                                 END_IF;
                               END_REGION PATH_DYNAMICS

                               REGION CIRCLE_PARAMETERS
                                 IF #statConfigCmdWords[#tempFollowValueCounter].%X4 THEN

                                   // Aux point
                                   FOR #tempCounter := 1 TO 3 DO
                                     IF #statParameterDefinition.followingValues[#tempFollowValueCounter].cmdParameters.circleParameters.auxPoint[#tempCounter] THEN
                                       // Set AuxPoint
                                       #tempParsedValues.cmdParameters.circleParameters.auxPoint[#tempCounter] := #tempParameterValue;
                                       #statParameterValid.cmdParameters.circleParameters.auxPoint[#tempCounter] := TRUE;
                                     END_IF;
                                   END_FOR;

                                   // PathChoice
                                   IF #statParameterDefinition.followingValues[#tempFollowValueCounter].cmdParameters.circleParameters.pathChoice THEN
                                     // Set PathChoice
                                     #tempParsedValues.cmdParameters.circleParameters.pathChoice := LREAL_TO_DINT(#tempParameterValue);
                                     #statParameterValid.cmdParameters.circleParameters.pathChoice := TRUE;
                                   END_IF;


                                   // CircMode
                                   IF #statParameterDefinition.followingValues[#tempFollowValueCounter].cmdParameters.circleParameters.circMode THEN
                                     // Set CircMode
                                     #tempParsedValues.cmdParameters.circleParameters.circMode := LREAL_TO_DINT(#tempParameterValue);
                                     #statParameterValid.cmdParameters.circleParameters.circMode := TRUE;
                                   END_IF;


                                   // CirclePlane
                                   IF #statParameterDefinition.followingValues[#tempFollowValueCounter].cmdParameters.circleParameters.circlePlane THEN
                                     // Set CirclePlane
                                     #tempParsedValues.cmdParameters.circleParameters.circlePlane := LREAL_TO_DINT(#tempParameterValue);
                                     #statParameterValid.cmdParameters.circleParameters.circlePlane := TRUE;
                                   END_IF;


                                   // Arc
                                   IF #statParameterDefinition.followingValues[#tempFollowValueCounter].cmdParameters.circleParameters.arc THEN
                                     // Set Arc
                                     #tempParsedValues.cmdParameters.circleParameters.arc := #tempParameterValue;
                                     #statParameterValid.cmdParameters.circleParameters.arc := TRUE;
                                   END_IF;


                                   // Radius
                                   IF #statParameterDefinition.followingValues[#tempFollowValueCounter].cmdParameters.circleParameters.radius THEN
                                     // Set Radius
                                     #tempParsedValues.cmdParameters.circleParameters.radius := #tempParameterValue;
                                     #statParameterValid.cmdParameters.circleParameters.radius := TRUE;
                                   END_IF;

                                 END_IF;
                               END_REGION CIRCLE_PARAMETERS

                               REGION BOOL_FLAGS
                                 // Always set first index of parsed values here
                                 // ----------------------------------------------------------------------------
                                 // Set Flags
                                 // ----------------------------------------------------------------------------
                                 IF #statParameterDefinition.followingValues[#tempFollowValueCounter].setFlags.flag THEN
                                   // Get parameter value
                                   #tempParsedValues.setFlags[1].flag := LREAL_TO_INT(#tempParameterValue);
                                   #statParameterValid.setFlags[1].flag := TRUE;
                                 END_IF;

                                 // ----------------------------------------------------------------------------
                                 // Flag Mode
                                 // ----------------------------------------------------------------------------
                                 IF #statParameterDefinition.followingValues[#tempFollowValueCounter].setFlags.flagMode THEN
                                   // Get parameter value
                                   #tempParsedValues.setFlags[1].flagMode := LREAL_TO_USINT(#tempParameterValue);
                                   #statParameterValid.setFlags[1].flagMode := TRUE;
                                 END_IF;


                                 // ----------------------------------------------------------------------------
                                 // Remaining Distance
                                 // ----------------------------------------------------------------------------
                                 IF #statParameterDefinition.followingValues[#tempFollowValueCounter].setFlags.remainingDistance THEN
                                   // Get parameter value
                                   #tempParsedValues.setFlags[1].remainingDistance := #tempParameterValue;
                                   #statParameterValid.setFlags[1].remainingDistance := TRUE;
                                 END_IF;

                               END_REGION BOOL_FLAGS

                               REGION LREAL_FLAGS
                                 // Always set first index of parsed values here
                                 // ----------------------------------------------------------------------------
                                 // Set Flags
                                 // ----------------------------------------------------------------------------
                                 IF #statParameterDefinition.followingValues[#tempFollowValueCounter].valueFlags.flag THEN
                                   // Get parameter value
                                   #tempParsedValues.valueFlags[1].flag := LREAL_TO_INT(#tempParameterValue);
                                   #statParameterValid.valueFlags[1].flag := TRUE;
                                 END_IF;

                                 // ----------------------------------------------------------------------------
                                 // Value
                                 // ----------------------------------------------------------------------------
                                 IF #statParameterDefinition.followingValues[#tempFollowValueCounter].valueFlags.value THEN
                                   // Get parameter value
                                   #tempParsedValues.valueFlags[1].value := #tempParameterValue;
                                   #statParameterValid.valueFlags[1].value := TRUE;
                                 END_IF;

                                 // ----------------------------------------------------------------------------
                                 // Flag Mode
                                 // ----------------------------------------------------------------------------
                                 IF #statParameterDefinition.followingValues[#tempFollowValueCounter].valueFlags.flagMode THEN
                                   // Get parameter value
                                   #tempParsedValues.valueFlags[1].flagMode := LREAL_TO_USINT(#tempParameterValue);
                                   #statParameterValid.valueFlags[1].flagMode := TRUE;
                                 END_IF;


                                 // ----------------------------------------------------------------------------
                                 // Remaining Distance
                                 // ----------------------------------------------------------------------------
                                 IF #statParameterDefinition.followingValues[#tempFollowValueCounter].valueFlags.remainingDistance THEN
                                   // Get parameter value
                                   #tempParsedValues.valueFlags[1].remainingDistance := #tempParameterValue;
                                   #statParameterValid.valueFlags[1].remainingDistance := TRUE;
                                 END_IF;

                               END_REGION LREAL_FLAGS

                             END_IF;
                           END_FOR;

                           // Exit loop in case of error
                           IF #statStatus.%X15 THEN
                             EXIT;
                           END_IF;
                         END_REGION GET_FOLLOW_VALUES   
                       END_IF;

                       IF #tempParseCounter = 2 THEN
                         REGION GET_DIRECT_VALUES
                           #tempCmdWord := #statDirectCmdWord;
                           #tempParsedValues := #statParameterDefinition.directValues;
                         END_REGION GET_DIRECT_VALUES
                       END_IF;


                       REGION SET_VALUES_IN_PATH_DATA_ELEMENT

                         IF #tempCmdWord.%X0 THEN

                           REGION CMD_TYPE
                             IF (#statParameterValid.cmdType AND #tempParseCounter = 1)
                               OR (NOT #statParameterValid.cmdType AND #tempParseCounter = 2)
                               AND #statParameterDefinition.priorities.cmdType > "LKINLANG_PRIO_UNRELEVANT"
                             THEN
                               // Get parameter value
                               #tempParameterValue := #tempParsedValues.cmdType;

                               // Set cmdType
                               #statPathDataValue.valueInt := #statActualCommand.pathDataElement.cmdType;
                               #statModalCmdValue.valueInt := #statModalCommand.pathDataElement.cmdType;
                               #statModalPrgValue.valueInt := #statModalProgram.pathDataElement.cmdType;

                               // Set value with follow val from above 
                               #tempReturnVal := "LKinLang_SetValue"(parameterValue := #tempParameterValue,
                                                                     parameterPriority := #statParameterDefinition.priorities.cmdType,
                                                                     validCountOfParameter := #statValidCounts.cmdType,
                                                                     parameterValueMin := -1,
                                                                     parameterValueMax := 100,
                                                                     properties := #statParameterDefinition.properties,
                                                                     errorString => #statErrorString,
                                                                     parameterCounter := #statElementCounter.cmdType,
                                                                     priorityCounter := #statActualCommand.priority.cmdType,
                                                                     modalCMDPrio := #statModalCommand.priority.cmdType,
                                                                     modalPRGPrio := #statModalProgram.priority.cmdType,
                                                                     parameterCounterInLine := #statElementCounterInLine.cmdType,
                                                                     pathDataValue := #statPathDataValue,
                                                                     modalCMDPathDataValue := #statModalCmdValue,
                                                                     modalPRGPathDataValue := #statModalPrgValue);

                               IF #tempReturnVal = 0 THEN
                                 #statActualCommand.pathDataElement.cmdType := #statPathDataValue.valueInt;
                                 #statModalCommand.pathDataElement.cmdType := #statModalCmdValue.valueInt;
                                 #statModalProgram.pathDataElement.cmdType := #statModalPrgValue.valueInt;
                               ELSE
                                 // Error
                                 #statStatus := #ERR_PARSING;
                                 #statErrorString := CONCAT(IN1 := #statErrorString, IN2 := '; Line: ');
                                 #statErrorString := CONCAT(IN1 := #statErrorString, IN2 := UDINT_TO_STRING(#statTokenizedLine.lineNo));
                                 EXIT;
                               END_IF;
                             END_IF;
                           END_REGION CMD_TYPE

                           REGION CMD_NAME
                             IF ((#statParameterValid.cmdName AND #tempParseCounter = 1)
                               OR (NOT #statParameterValid.cmdName AND #tempParseCounter = 2))
                               AND #tempParsedValues.cmdName <> ''
                               AND #statParameterDefinition.priorities.cmdName > "LKINLANG_PRIO_UNRELEVANT"
                             THEN

                               // Get parameter value
                               #tempParameterValue := STRING_TO_INT(#tempParsedValues.cmdName);

                               // Set cmdName
                               #statPathDataValue.valueInt := STRING_TO_INT(#statActualCommand.pathDataElement.cmdName);
                               #statModalCmdValue.valueInt := STRING_TO_INT(#statModalCommand.pathDataElement.cmdName);
                               #statModalPrgValue.valueInt := STRING_TO_INT(#statModalProgram.pathDataElement.cmdName);

                               // Set value with follow val from above 
                               #tempReturnVal := "LKinLang_SetValue"(parameterValue := #tempParameterValue,
                                                                     parameterPriority := #statParameterDefinition.priorities.cmdName,
                                                                     validCountOfParameter := #statValidCounts.cmdName,
                                                                     parameterValueMin := #MINVAL_INT,
                                                                     parameterValueMax := #MAXVAL_INT,
                                                                     properties := #statParameterDefinition.properties,
                                                                     errorString => #statErrorString,
                                                                     parameterCounter := #statElementCounter.cmdName,
                                                                     priorityCounter := #statActualCommand.priority.cmdName,
                                                                     modalCMDPrio := #statModalCommand.priority.cmdName,
                                                                     modalPRGPrio := #statModalProgram.priority.cmdName,
                                                                     parameterCounterInLine := #statElementCounterInLine.cmdName,
                                                                     pathDataValue := #statPathDataValue,
                                                                     modalCMDPathDataValue := #statModalCmdValue,
                                                                     modalPRGPathDataValue := #statModalPrgValue);

                               IF #tempReturnVal = 0 THEN
                                 #statActualCommand.pathDataElement.cmdName := INT_TO_STRING(#statPathDataValue.valueInt);

                                 // 16.07.2019 FR: Delete "+" sign from string
                                 IF #statPathDataValue.valueInt >= 0.0 THEN
                                   #statActualCommand.pathDataElement.cmdName := DELETE(IN := #statActualCommand.pathDataElement.cmdName, L := 1, P := 1);
                                 ELSE
                                   ; // Keep "-" sign
                                 END_IF;

                                 #statModalCommand.pathDataElement.cmdName := INT_TO_STRING(#statModalCmdValue.valueInt);
                                 #statModalProgram.pathDataElement.cmdName := INT_TO_STRING(#statModalPrgValue.valueInt);
                               ELSE
                                 // Error
                                 #statStatus := #ERR_PARSING;
                                 #statErrorString := CONCAT(IN1 := #statErrorString, IN2 := '; Line: ');
                                 #statErrorString := CONCAT(IN1 := #statErrorString, IN2 := UDINT_TO_STRING(#statTokenizedLine.lineNo));
                                 EXIT;
                               END_IF;
                             END_IF;
                           END_REGION CMD_NAME

                           REGION COORDINATES
                             IF #tempCmdWord.%X1 THEN // Coordinates are set

                               // X coordinate
                               IF (#statParameterValid.cmdCoordinates.cartesianPosition.x AND #tempParseCounter = 1)
                                 OR (NOT #statParameterValid.cmdCoordinates.cartesianPosition.x AND #tempParseCounter = 2)
                                 AND #statParameterDefinition.priorities.cmdCoordinates.cartesianPosition.x > "LKINLANG_PRIO_UNRELEVANT"
                               THEN

                                 // Get parameter value
                                 #tempParameterValue := #tempParsedValues.cmdCoordinates.cartesianPosition.x;

                                 // Set X
                                 #statPathDataValue.valueLReal := #statActualCommand.pathDataElement.cmdCoordinates.cartesianPosition.x;
                                 #statModalCmdValue.valueLReal := #statModalCommand.pathDataElement.cmdCoordinates.cartesianPosition.x;
                                 #statModalPrgValue.valueLReal := #statModalProgram.pathDataElement.cmdCoordinates.cartesianPosition.x;

                                 // Set value with follow val from above 
                                 #tempReturnVal := "LKinLang_SetValue"(parameterValue := #tempParameterValue,
                                                                       parameterPriority := #statParameterDefinition.priorities.cmdCoordinates.cartesianPosition.x,
                                                                       validCountOfParameter := #statValidCounts.cmdCoordinates.cartesianPosition.x,
                                                                       parameterValueMin := #MINVAL_LREAL,
                                                                       parameterValueMax := #MAXVAL_LREAL,
                                                                       properties := #statParameterDefinition.properties,
                                                                       errorString => #statErrorString,
                                                                       parameterCounter := #statElementCounter.cmdCoordinates.cartesianPosition.x,
                                                                       priorityCounter := #statActualCommand.priority.cmdCoordinates.cartesianPosition.x,
                                                                       modalCMDPrio := #statModalCommand.priority.cmdCoordinates.cartesianPosition.x,
                                                                       modalPRGPrio := #statModalProgram.priority.cmdCoordinates.cartesianPosition.x,
                                                                       parameterCounterInLine := #statElementCounterInLine.cmdCoordinates.cartesianPosition.x,
                                                                       pathDataValue := #statPathDataValue,
                                                                       modalCMDPathDataValue := #statModalCmdValue,
                                                                       modalPRGPathDataValue := #statModalPrgValue);

                                 IF #tempReturnVal = 0 THEN
                                   #statActualCommand.pathDataElement.cmdCoordinates.cartesianPosition.x := #statPathDataValue.valueLReal;
                                   #statModalCommand.pathDataElement.cmdCoordinates.cartesianPosition.x := #statModalCmdValue.valueLReal;
                                   #statModalProgram.pathDataElement.cmdCoordinates.cartesianPosition.x := #statModalPrgValue.valueLReal;

                                   // Set parameter valid bit for MovePath 
                                   #statActualCommand.pathDataElement.parameterValid[1] := TRUE;
                                 ELSE
                                   // Error
                                   #statStatus := #ERR_PARSING;
                                   #statErrorString := CONCAT(IN1 := #statErrorString, IN2 := '; Line: ');
                                   #statErrorString := CONCAT(IN1 := #statErrorString, IN2 := UDINT_TO_STRING(#statTokenizedLine.lineNo));
                                   EXIT;
                                 END_IF;
                               END_IF;


                               // Y coordinate
                               IF (#statParameterValid.cmdCoordinates.cartesianPosition.y AND #tempParseCounter = 1)
                                 OR (NOT #statParameterValid.cmdCoordinates.cartesianPosition.y AND #tempParseCounter = 2)
                                 AND #statParameterDefinition.priorities.cmdCoordinates.cartesianPosition.y > "LKINLANG_PRIO_UNRELEVANT"
                               THEN

                                 // Get parameter value
                                 #tempParameterValue := #tempParsedValues.cmdCoordinates.cartesianPosition.y;

                                 // Set Y
                                 #statPathDataValue.valueLReal := #statActualCommand.pathDataElement.cmdCoordinates.cartesianPosition.y;
                                 #statModalCmdValue.valueLReal := #statModalCommand.pathDataElement.cmdCoordinates.cartesianPosition.y;
                                 #statModalPrgValue.valueLReal := #statModalProgram.pathDataElement.cmdCoordinates.cartesianPosition.y;

                                 // Set value with follow val from above 
                                 #tempReturnVal := "LKinLang_SetValue"(parameterValue := #tempParameterValue,
                                                                       parameterPriority := #statParameterDefinition.priorities.cmdCoordinates.cartesianPosition.y,
                                                                       validCountOfParameter := #statValidCounts.cmdCoordinates.cartesianPosition.y,
                                                                       parameterValueMin := #MINVAL_LREAL,
                                                                       parameterValueMax := #MAXVAL_LREAL,
                                                                       properties := #statParameterDefinition.properties,
                                                                       errorString => #statErrorString,
                                                                       parameterCounter := #statElementCounter.cmdCoordinates.cartesianPosition.y,
                                                                       priorityCounter := #statActualCommand.priority.cmdCoordinates.cartesianPosition.y,
                                                                       modalCMDPrio := #statModalCommand.priority.cmdCoordinates.cartesianPosition.y,
                                                                       modalPRGPrio := #statModalProgram.priority.cmdCoordinates.cartesianPosition.y,
                                                                       parameterCounterInLine := #statElementCounterInLine.cmdCoordinates.cartesianPosition.y,
                                                                       pathDataValue := #statPathDataValue,
                                                                       modalCMDPathDataValue := #statModalCmdValue,
                                                                       modalPRGPathDataValue := #statModalPrgValue);

                                 IF #tempReturnVal = 0 THEN
                                   #statActualCommand.pathDataElement.cmdCoordinates.cartesianPosition.y := #statPathDataValue.valueLReal;
                                   #statModalCommand.pathDataElement.cmdCoordinates.cartesianPosition.y := #statModalCmdValue.valueLReal;
                                   #statModalProgram.pathDataElement.cmdCoordinates.cartesianPosition.y := #statModalPrgValue.valueLReal;

                                   // Set parameter valid bit for MovePath 
                                   #statActualCommand.pathDataElement.parameterValid[2] := TRUE;
                                 ELSE
                                   // Error
                                   #statStatus := #ERR_PARSING;
                                   #statErrorString := CONCAT(IN1 := #statErrorString, IN2 := '; Line: ');
                                   #statErrorString := CONCAT(IN1 := #statErrorString, IN2 := UDINT_TO_STRING(#statTokenizedLine.lineNo));
                                   EXIT;
                                 END_IF;
                               END_IF;



                               // Z coordinate
                               IF (#statParameterValid.cmdCoordinates.cartesianPosition.z AND #tempParseCounter = 1)
                                 OR (NOT #statParameterValid.cmdCoordinates.cartesianPosition.z AND #tempParseCounter = 2)
                                 AND #statParameterDefinition.priorities.cmdCoordinates.cartesianPosition.z > "LKINLANG_PRIO_UNRELEVANT"
                               THEN

                                 // Get parameter value
                                 #tempParameterValue := #tempParsedValues.cmdCoordinates.cartesianPosition.z;

                                 // Set Z
                                 #statPathDataValue.valueLReal := #statActualCommand.pathDataElement.cmdCoordinates.cartesianPosition.z;
                                 #statModalCmdValue.valueLReal := #statModalCommand.pathDataElement.cmdCoordinates.cartesianPosition.z;
                                 #statModalPrgValue.valueLReal := #statModalProgram.pathDataElement.cmdCoordinates.cartesianPosition.z;

                                 // Set value with follow val from above 
                                 #tempReturnVal := "LKinLang_SetValue"(parameterValue := #tempParameterValue,
                                                                       parameterPriority := #statParameterDefinition.priorities.cmdCoordinates.cartesianPosition.z,
                                                                       validCountOfParameter := #statValidCounts.cmdCoordinates.cartesianPosition.z,
                                                                       parameterValueMin := #MINVAL_LREAL,
                                                                       parameterValueMax := #MAXVAL_LREAL,
                                                                       properties := #statParameterDefinition.properties,
                                                                       errorString => #statErrorString,
                                                                       parameterCounter := #statElementCounter.cmdCoordinates.cartesianPosition.z,
                                                                       priorityCounter := #statActualCommand.priority.cmdCoordinates.cartesianPosition.z,
                                                                       modalCMDPrio := #statModalCommand.priority.cmdCoordinates.cartesianPosition.z,
                                                                       modalPRGPrio := #statModalProgram.priority.cmdCoordinates.cartesianPosition.z,
                                                                       parameterCounterInLine := #statElementCounterInLine.cmdCoordinates.cartesianPosition.z,
                                                                       pathDataValue := #statPathDataValue,
                                                                       modalCMDPathDataValue := #statModalCmdValue,
                                                                       modalPRGPathDataValue := #statModalPrgValue);

                                 IF #tempReturnVal = 0 THEN
                                   #statActualCommand.pathDataElement.cmdCoordinates.cartesianPosition.z := #statPathDataValue.valueLReal;
                                   #statModalCommand.pathDataElement.cmdCoordinates.cartesianPosition.z := #statModalCmdValue.valueLReal;
                                   #statModalProgram.pathDataElement.cmdCoordinates.cartesianPosition.z := #statModalPrgValue.valueLReal;

                                   // Set parameter valid bit for MovePath 
                                   #statActualCommand.pathDataElement.parameterValid[3] := TRUE;
                                 ELSE
                                   // Error
                                   #statStatus := #ERR_PARSING;
                                   #statErrorString := CONCAT(IN1 := #statErrorString, IN2 := '; Line: ');
                                   #statErrorString := CONCAT(IN1 := #statErrorString, IN2 := UDINT_TO_STRING(#statTokenizedLine.lineNo));
                                   EXIT;
                                 END_IF;
                               END_IF;


                               // A coordinate
                               IF (#statParameterValid.cmdCoordinates.cartesianPosition.a AND #tempParseCounter = 1)
                                 OR (NOT #statParameterValid.cmdCoordinates.cartesianPosition.a AND #tempParseCounter = 2)
                                 AND #statParameterDefinition.priorities.cmdCoordinates.cartesianPosition.a > "LKINLANG_PRIO_UNRELEVANT"
                               THEN

                                 // Get parameter value
                                 #tempParameterValue := #tempParsedValues.cmdCoordinates.cartesianPosition.a;

                                 // Set A
                                 #statPathDataValue.valueLReal := #statActualCommand.pathDataElement.cmdCoordinates.cartesianPosition.a;
                                 #statModalCmdValue.valueLReal := #statModalCommand.pathDataElement.cmdCoordinates.cartesianPosition.a;
                                 #statModalPrgValue.valueLReal := #statModalProgram.pathDataElement.cmdCoordinates.cartesianPosition.a;

                                 // Set value with follow val from above 
                                 #tempReturnVal := "LKinLang_SetValue"(parameterValue := #tempParameterValue,
                                                                       parameterPriority := #statParameterDefinition.priorities.cmdCoordinates.cartesianPosition.a,
                                                                       validCountOfParameter := #statValidCounts.cmdCoordinates.cartesianPosition.a,
                                                                       parameterValueMin := #MINVAL_LREAL,
                                                                       parameterValueMax := #MAXVAL_LREAL,
                                                                       properties := #statParameterDefinition.properties,
                                                                       errorString => #statErrorString,
                                                                       parameterCounter := #statElementCounter.cmdCoordinates.cartesianPosition.a,
                                                                       priorityCounter := #statActualCommand.priority.cmdCoordinates.cartesianPosition.a,
                                                                       modalCMDPrio := #statModalCommand.priority.cmdCoordinates.cartesianPosition.a,
                                                                       modalPRGPrio := #statModalProgram.priority.cmdCoordinates.cartesianPosition.a,
                                                                       parameterCounterInLine := #statElementCounterInLine.cmdCoordinates.cartesianPosition.a,
                                                                       pathDataValue := #statPathDataValue,
                                                                       modalCMDPathDataValue := #statModalCmdValue,
                                                                       modalPRGPathDataValue := #statModalPrgValue);

                                 IF #tempReturnVal = 0 THEN
                                   #statActualCommand.pathDataElement.cmdCoordinates.cartesianPosition.a := #statPathDataValue.valueLReal;
                                   #statModalCommand.pathDataElement.cmdCoordinates.cartesianPosition.a := #statModalCmdValue.valueLReal;
                                   #statModalProgram.pathDataElement.cmdCoordinates.cartesianPosition.a := #statModalPrgValue.valueLReal;

                                   // Set parameter valid bit for MovePath 
                                   #statActualCommand.pathDataElement.parameterValid[4] := TRUE;
                                 ELSE
                                   // Error
                                   #statStatus := #ERR_PARSING;
                                   #statErrorString := CONCAT(IN1 := #statErrorString, IN2 := '; Line: ');
                                   #statErrorString := CONCAT(IN1 := #statErrorString, IN2 := UDINT_TO_STRING(#statTokenizedLine.lineNo));
                                   EXIT;
                                 END_IF;
                               END_IF;


                               // CoordSystem coordinate
                               IF (#statParameterValid.cmdCoordinates.coordSystem AND #tempParseCounter = 1)
                                 OR (NOT #statParameterValid.cmdCoordinates.coordSystem AND #tempParseCounter = 2)
                                 AND #statParameterDefinition.priorities.cmdCoordinates.coordSystem > "LKINLANG_PRIO_UNRELEVANT"
                               THEN

                                 // Get parameter value
                                 #tempParameterValue := #tempParsedValues.cmdCoordinates.coordSystem;

                                 // Set CS
                                 #statPathDataValue.valueDint := #statActualCommand.pathDataElement.cmdCoordinates.coordSystem;
                                 #statModalCmdValue.valueDint := #statModalCommand.pathDataElement.cmdCoordinates.coordSystem;
                                 #statModalPrgValue.valueDint := #statModalProgram.pathDataElement.cmdCoordinates.coordSystem;

                                 // Set value with follow val from above 
                                 #tempReturnVal := "LKinLang_SetValue"(parameterValue := #tempParameterValue,
                                                                       parameterPriority := #statParameterDefinition.priorities.cmdCoordinates.coordSystem,
                                                                       validCountOfParameter := #statValidCounts.cmdCoordinates.coordSystem,
                                                                       parameterValueMin := 0,
                                                                       parameterValueMax := 3,
                                                                       properties := #statParameterDefinition.properties,
                                                                       errorString => #statErrorString,
                                                                       parameterCounter := #statElementCounter.cmdCoordinates.coordSystem,
                                                                       priorityCounter := #statActualCommand.priority.cmdCoordinates.coordSystem,
                                                                       modalCMDPrio := #statModalCommand.priority.cmdCoordinates.coordSystem,
                                                                       modalPRGPrio := #statModalProgram.priority.cmdCoordinates.coordSystem,
                                                                       parameterCounterInLine := #statElementCounterInLine.cmdCoordinates.coordSystem,
                                                                       pathDataValue := #statPathDataValue,
                                                                       modalCMDPathDataValue := #statModalCmdValue,
                                                                       modalPRGPathDataValue := #statModalPrgValue);

                                 IF #tempReturnVal = 0 THEN
                                   #statActualCommand.pathDataElement.cmdCoordinates.coordSystem := #statPathDataValue.valueDint;
                                   #statModalCommand.pathDataElement.cmdCoordinates.coordSystem := #statModalCmdValue.valueDint;
                                   #statModalProgram.pathDataElement.cmdCoordinates.coordSystem := #statModalPrgValue.valueDint;
                                 ELSE
                                   // Error
                                   #statStatus := #ERR_PARSING;
                                   #statErrorString := CONCAT(IN1 := #statErrorString, IN2 := '; Line: ');
                                   #statErrorString := CONCAT(IN1 := #statErrorString, IN2 := UDINT_TO_STRING(#statTokenizedLine.lineNo));
                                   EXIT;
                                 END_IF;
                               END_IF;

                             END_IF;
                           END_REGION COORDINATES

                           REGION CMD_PARAMETERS

                             IF #tempCmdWord.%X2 THEN // Parameter are to be set

                               REGION GENERAL_PARAMETERS

                                 // Buffer mode
                                 IF (#statParameterValid.cmdParameters.bufferMode AND #tempParseCounter = 1)
                                   OR (NOT #statParameterValid.cmdParameters.bufferMode AND #tempParseCounter = 2)
                                   AND #statParameterDefinition.priorities.cmdParameters.bufferMode > "LKINLANG_PRIO_UNRELEVANT"
                                 THEN

                                   // Get parameter value
                                   #tempParameterValue := #tempParsedValues.cmdParameters.bufferMode;

                                   // Set Velocity
                                   #statPathDataValue.valueDint := #statActualCommand.pathDataElement.cmdParameters.bufferMode;
                                   #statModalCmdValue.valueDint := #statModalCommand.pathDataElement.cmdParameters.bufferMode;
                                   #statModalPrgValue.valueDint := #statModalProgram.pathDataElement.cmdParameters.bufferMode;

                                   // Set value with follow val from above 
                                   #tempReturnVal := "LKinLang_SetValue"(parameterValue := #tempParameterValue,
                                                                         parameterPriority := #statParameterDefinition.priorities.cmdParameters.bufferMode,
                                                                         validCountOfParameter := #statValidCounts.cmdParameters.bufferMode,
                                                                         parameterValueMin := 1,
                                                                         parameterValueMax := 5,
                                                                         properties := #statParameterDefinition.properties,
                                                                         errorString => #statErrorString,
                                                                         parameterCounter := #statElementCounter.cmdParameters.bufferMode,
                                                                         priorityCounter := #statActualCommand.priority.cmdParameters.bufferMode,
                                                                         modalCMDPrio := #statModalCommand.priority.cmdParameters.bufferMode,
                                                                         modalPRGPrio := #statModalProgram.priority.cmdParameters.bufferMode,
                                                                         parameterCounterInLine := #statElementCounterInLine.cmdParameters.bufferMode,
                                                                         pathDataValue := #statPathDataValue,
                                                                         modalCMDPathDataValue := #statModalCmdValue,
                                                                         modalPRGPathDataValue := #statModalPrgValue);

                                   IF #tempReturnVal = 0 THEN
                                     #statActualCommand.pathDataElement.cmdParameters.bufferMode := #statPathDataValue.valueDint;
                                     #statModalCommand.pathDataElement.cmdParameters.bufferMode := #statModalCmdValue.valueDint;
                                     #statModalProgram.pathDataElement.cmdParameters.bufferMode := #statModalPrgValue.valueDint;
                                   ELSE
                                     // Error
                                     #statStatus := #ERR_PARSING;
                                     #statErrorString := CONCAT(IN1 := #statErrorString, IN2 := '; Line: ');
                                     #statErrorString := CONCAT(IN1 := #statErrorString, IN2 := UDINT_TO_STRING(#statTokenizedLine.lineNo));
                                     EXIT;
                                   END_IF;
                                 END_IF;

                                 // Dynamic adaption
                                 IF (#statParameterValid.cmdParameters.dynamicAdaption AND #tempParseCounter = 1)
                                   OR (NOT #statParameterValid.cmdParameters.dynamicAdaption AND #tempParseCounter = 2)
                                   AND #statParameterDefinition.priorities.cmdParameters.dynamicAdaption > "LKINLANG_PRIO_UNRELEVANT"
                                 THEN

                                   // Get parameter value
                                   #tempParameterValue := #tempParsedValues.cmdParameters.dynamicAdaption;

                                   // Set Velocity
                                   #statPathDataValue.valueDint := #statActualCommand.pathDataElement.cmdParameters.dynamicAdaption;
                                   #statModalCmdValue.valueDint := #statModalCommand.pathDataElement.cmdParameters.dynamicAdaption;
                                   #statModalPrgValue.valueDint := #statModalProgram.pathDataElement.cmdParameters.dynamicAdaption;

                                   // Set value with follow val from above 
                                   #tempReturnVal := "LKinLang_SetValue"(parameterValue := #tempParameterValue,
                                                                         parameterPriority := #statParameterDefinition.priorities.cmdParameters.dynamicAdaption,
                                                                         validCountOfParameter := #statValidCounts.cmdParameters.dynamicAdaption,
                                                                         parameterValueMin := -1,
                                                                         parameterValueMax := 2,
                                                                         properties := #statParameterDefinition.properties,
                                                                         errorString => #statErrorString,
                                                                         parameterCounter := #statElementCounter.cmdParameters.dynamicAdaption,
                                                                         priorityCounter := #statActualCommand.priority.cmdParameters.dynamicAdaption,
                                                                         modalCMDPrio := #statModalCommand.priority.cmdParameters.dynamicAdaption,
                                                                         modalPRGPrio := #statModalProgram.priority.cmdParameters.dynamicAdaption,
                                                                         parameterCounterInLine := #statElementCounterInLine.cmdParameters.dynamicAdaption,
                                                                         pathDataValue := #statPathDataValue,
                                                                         modalCMDPathDataValue := #statModalCmdValue,
                                                                         modalPRGPathDataValue := #statModalPrgValue);

                                   IF #tempReturnVal = 0 THEN
                                     #statActualCommand.pathDataElement.cmdParameters.dynamicAdaption := #statPathDataValue.valueDint;
                                     #statModalCommand.pathDataElement.cmdParameters.dynamicAdaption := #statModalCmdValue.valueDint;
                                     #statModalProgram.pathDataElement.cmdParameters.dynamicAdaption := #statModalPrgValue.valueDint;
                                   ELSE
                                     // Error
                                     #statStatus := #ERR_PARSING;
                                     #statErrorString := CONCAT(IN1 := #statErrorString, IN2 := '; Line: ');
                                     #statErrorString := CONCAT(IN1 := #statErrorString, IN2 := UDINT_TO_STRING(#statTokenizedLine.lineNo));
                                     EXIT;
                                   END_IF;
                                 END_IF;

                                 // Offset Parameter
                                 // Offset Parameter number
                                 IF (#statParameterValid.cmdParameters.offsetParameters.offsetParaNo AND #tempParseCounter = 1)
                                   OR (NOT #statParameterValid.cmdParameters.offsetParameters.offsetParaNo AND #tempParseCounter = 2)
                                   AND #statParameterDefinition.priorities.cmdParameters.offsetParameters.offsetParaNo > "LKINLANG_PRIO_UNRELEVANT"
                                 THEN

                                   // Get parameter value
                                   #tempParameterValue := #tempParsedValues.cmdParameters.offsetParameters.offsetParaNo;

                                   // Set Velocity
                                   #statPathDataValue.valueDint := #statActualCommand.pathDataElement.cmdParameters.offsetParameters.offsetParaNo;
                                   #statModalCmdValue.valueDint := #statModalCommand.pathDataElement.cmdParameters.offsetParameters.offsetParaNo;
                                   #statModalPrgValue.valueDint := #statModalProgram.pathDataElement.cmdParameters.offsetParameters.offsetParaNo;

                                   // Set value with follow val from above 
                                   #tempReturnVal := "LKinLang_SetValue"(parameterValue := #tempParameterValue,
                                                                         parameterPriority := #statParameterDefinition.priorities.cmdParameters.offsetParameters.offsetParaNo,
                                                                         validCountOfParameter := #statValidCounts.cmdParameters.offsetParameters.offsetParaNo,
                                                                         parameterValueMin := -1,
                                                                         parameterValueMax := #MAXVAL_INT,
                                                                         properties := #statParameterDefinition.properties,
                                                                         errorString => #statErrorString,
                                                                         parameterCounter := #statElementCounter.cmdParameters.offsetParameters.offsetParaNo,
                                                                         priorityCounter := #statActualCommand.priority.cmdParameters.offsetParameters.offsetParaNo,
                                                                         modalCMDPrio := #statModalCommand.priority.cmdParameters.offsetParameters.offsetParaNo,
                                                                         modalPRGPrio := #statModalProgram.priority.cmdParameters.offsetParameters.offsetParaNo,
                                                                         parameterCounterInLine := #statElementCounterInLine.cmdParameters.offsetParameters.offsetParaNo,
                                                                         pathDataValue := #statPathDataValue,
                                                                         modalCMDPathDataValue := #statModalCmdValue,
                                                                         modalPRGPathDataValue := #statModalPrgValue);

                                   IF #tempReturnVal = 0 THEN
                                     #statActualCommand.pathDataElement.cmdParameters.offsetParameters.offsetParaNo := #statPathDataValue.valueInt;
                                     #statModalCommand.pathDataElement.cmdParameters.offsetParameters.offsetParaNo := #statModalCmdValue.valueInt;
                                     #statModalProgram.pathDataElement.cmdParameters.offsetParameters.offsetParaNo := #statModalPrgValue.valueInt;
                                   ELSE
                                     // Error
                                     #statStatus := #ERR_PARSING;
                                     #statErrorString := CONCAT(IN1 := #statErrorString, IN2 := '; Line: ');
                                     #statErrorString := CONCAT(IN1 := #statErrorString, IN2 := UDINT_TO_STRING(#statTokenizedLine.lineNo));
                                     EXIT;
                                   END_IF;
                                 END_IF;

                                 // Offset Main Path plane
                                 IF (#statParameterValid.cmdParameters.offsetParameters.mainPathPlane AND #tempParseCounter = 1)
                                   OR (NOT #statParameterValid.cmdParameters.offsetParameters.mainPathPlane AND #tempParseCounter = 2)
                                   AND #statParameterDefinition.priorities.cmdParameters.offsetParameters.mainPathPlane > "LKINLANG_PRIO_UNRELEVANT"
                                 THEN

                                   // Get parameter value
                                   #tempParameterValue := #tempParsedValues.cmdParameters.offsetParameters.mainPathPlane;

                                   // Set Velocity
                                   #statPathDataValue.valueDint := #statActualCommand.pathDataElement.cmdParameters.offsetParameters.mainPathPlane;
                                   #statModalCmdValue.valueDint := #statModalCommand.pathDataElement.cmdParameters.offsetParameters.mainPathPlane;
                                   #statModalPrgValue.valueDint := #statModalProgram.pathDataElement.cmdParameters.offsetParameters.mainPathPlane;

                                   // Set value with follow val from above 
                                   #tempReturnVal := "LKinLang_SetValue"(parameterValue := #tempParameterValue,
                                                                         parameterPriority := #statParameterDefinition.priorities.cmdParameters.offsetParameters.mainPathPlane,
                                                                         validCountOfParameter := #statValidCounts.cmdParameters.offsetParameters.mainPathPlane,
                                                                         parameterValueMin := 0,
                                                                         parameterValueMax := 2,
                                                                         properties := #statParameterDefinition.properties,
                                                                         errorString => #statErrorString,
                                                                         parameterCounter := #statElementCounter.cmdParameters.offsetParameters.mainPathPlane,
                                                                         priorityCounter := #statActualCommand.priority.cmdParameters.offsetParameters.mainPathPlane,
                                                                         modalCMDPrio := #statModalCommand.priority.cmdParameters.offsetParameters.mainPathPlane,
                                                                         modalPRGPrio := #statModalProgram.priority.cmdParameters.offsetParameters.mainPathPlane,
                                                                         parameterCounterInLine := #statElementCounterInLine.cmdParameters.offsetParameters.mainPathPlane,
                                                                         pathDataValue := #statPathDataValue,
                                                                         modalCMDPathDataValue := #statModalCmdValue,
                                                                         modalPRGPathDataValue := #statModalPrgValue);

                                   IF #tempReturnVal = 0 THEN
                                     #statActualCommand.pathDataElement.cmdParameters.offsetParameters.mainPathPlane := #statPathDataValue.valueInt;
                                     #statModalCommand.pathDataElement.cmdParameters.offsetParameters.mainPathPlane := #statModalCmdValue.valueInt;
                                     #statModalProgram.pathDataElement.cmdParameters.offsetParameters.mainPathPlane := #statModalPrgValue.valueInt;
                                   ELSE
                                     // Error
                                     #statStatus := #ERR_PARSING;
                                     #statErrorString := CONCAT(IN1 := #statErrorString, IN2 := '; Line: ');
                                     #statErrorString := CONCAT(IN1 := #statErrorString, IN2 := UDINT_TO_STRING(#statTokenizedLine.lineNo));
                                     EXIT;
                                   END_IF;
                                 END_IF;

                                 // Transition parameter
                                 FOR #tempCounter := 1 TO 5 DO
                                   IF (#statParameterValid.cmdParameters.transitionParameters[#tempCounter] AND #tempParseCounter = 1)
                                     OR (NOT #statParameterValid.cmdParameters.transitionParameters[#tempCounter] AND #tempParseCounter = 2)
                                     AND #statParameterDefinition.priorities.cmdParameters.transitionParameters[#tempCounter] > "LKINLANG_PRIO_UNRELEVANT"
                                   THEN

                                     // Get parameter value
                                     #tempParameterValue := #tempParsedValues.cmdParameters.transitionParameters[#tempCounter];

                                     // Set Velocity
                                     #statPathDataValue.valueLReal := #statActualCommand.pathDataElement.cmdParameters.transitionParameters[#tempCounter];
                                     #statModalCmdValue.valueLReal := #statModalCommand.pathDataElement.cmdParameters.transitionParameters[#tempCounter];
                                     #statModalPrgValue.valueLReal := #statModalProgram.pathDataElement.cmdParameters.transitionParameters[#tempCounter];

                                     // Set value with follow val from above 
                                     #tempReturnVal := "LKinLang_SetValue"(parameterValue := #tempParameterValue,
                                                                           parameterPriority := #statParameterDefinition.priorities.cmdParameters.transitionParameters[#tempCounter],
                                                                           validCountOfParameter := #statValidCounts.cmdParameters.transitionParameters[#tempCounter],
                                                                           parameterValueMin := #MINVAL_LREAL,
                                                                           parameterValueMax := #MAXVAL_LREAL,
                                                                           properties := #statParameterDefinition.properties,
                                                                           errorString => #statErrorString,
                                                                           parameterCounter := #statElementCounter.cmdParameters.transitionParameters[#tempCounter],
                                                                           priorityCounter := #statActualCommand.priority.cmdParameters.transitionParameters[#tempCounter],
                                                                           modalCMDPrio := #statModalCommand.priority.cmdParameters.transitionParameters[#tempCounter],
                                                                           modalPRGPrio := #statModalProgram.priority.cmdParameters.transitionParameters[#tempCounter],
                                                                           parameterCounterInLine := #statElementCounterInLine.cmdParameters.transitionParameters[#tempCounter],
                                                                           pathDataValue := #statPathDataValue,
                                                                           modalCMDPathDataValue := #statModalCmdValue,
                                                                           modalPRGPathDataValue := #statModalPrgValue);

                                     IF #tempReturnVal = 0 THEN
                                       #statActualCommand.pathDataElement.cmdParameters.transitionParameters[#tempCounter] := #statPathDataValue.valueLReal;
                                       #statModalCommand.pathDataElement.cmdParameters.transitionParameters[#tempCounter] := #statModalCmdValue.valueLReal;
                                       #statModalProgram.pathDataElement.cmdParameters.transitionParameters[#tempCounter] := #statModalPrgValue.valueLReal;
                                     ELSE
                                       // Error
                                       #statStatus := #ERR_PARSING;
                                       #statErrorString := CONCAT(IN1 := #statErrorString, IN2 := '; Line: ');
                                       #statErrorString := CONCAT(IN1 := #statErrorString, IN2 := UDINT_TO_STRING(#statTokenizedLine.lineNo));
                                       EXIT;
                                     END_IF;
                                   END_IF;
                                 END_FOR;

                               END_REGION GENERAL_PARAMETERS

                               REGION PATH_DYNAMICS
                                 IF #tempCmdWord.%X3 THEN // Dynamics are to be set

                                   // Velocity
                                   IF (#statParameterValid.cmdParameters.pathDynamics.velocity AND #tempParseCounter = 1)
                                     OR (NOT #statParameterValid.cmdParameters.pathDynamics.velocity AND #tempParseCounter = 2)
                                     AND #statParameterDefinition.priorities.cmdParameters.pathDynamics.velocity > "LKINLANG_PRIO_UNRELEVANT"
                                   THEN


                                     // Check for wait time only whe velocity is trying to be set 01.02.2019
                                     // Testing non modal F for wait time 24.01.2019
                                     REGION CHECK_FOR_WAIT_TIME
                                       // Pre check for wait time 
                                       FOR #tempWaitCheckCounter := 1 TO #statTokenizedLine.numberOfToken BY 1 DO
                                         //#statWaitParameterDef := #statParameterDefEmpty;
                                         #statTokenCheck.actual := #statTokenizedLine.lineToken[#tempWaitCheckCounter];

                                         //Get previous token
                                         IF #tempWaitCheckCounter > 1 THEN
                                           #statTokenCheck.previous := #statTokenizedLine.lineToken[#tempWaitCheckCounter - 1];
                                         ELSE
                                           #statTokenCheck.previous := '';
                                         END_IF;

                                         // Only check token for parameter if it is a letter --> numeric is skipped
                                         IF STRING_TO_LREAL(#statTokenCheck.actual) = 0.0 THEN

                                           // Testing 28.01.2019
                                           // Old parameter def
                                           #tempParameterIndex := "LKinLang_IsTokenParameter"(tokenToCheck := #statTokenCheck,
                                                                                              language := #language,
                                                                                              lastIndexLookUp := #statLastIndexLookUp,
                                                                                              parameterDefinition := #tempWaitParameterDefinition,
                                                                                              parameterLookUpTable := #statParameterLookUpTable,
                                                                                              parameterDefaults := #parameterDefaults,
                                                                                              directCmdWord := #statDirectCmdWord,
                                                                                              configCmdWords := #statConfigCmdWords);

                                           // Check direct value, also check follow value ?
                                           // What about modal value ?
                                           IF #tempWaitParameterDefinition.directValues.cmdType = 100 THEN
                                             #tempWaitTime := TRUE; // Use this variable later on to reset modal properties when setting velocity parameter
                                             EXIT;
                                           END_IF;

                                         END_IF;
                                       END_FOR;
                                     END_REGION CHECK_FOR_WAIT_TIME

                                     // Testing 24.01.2019 
                                     // Reset modal when wait time is set
                                     IF #tempWaitTime THEN
                                       ;
                                       #statParameterDefinition.properties := #statParameterDefinition.properties AND NOT "LKINLANG_PRG_MODAL";
                                     ELSE
                                       ; // Do not change property
                                     END_IF;


                                     // Get parameter value
                                     #tempParameterValue := #tempParsedValues.cmdParameters.pathDynamics.velocity;

                                     // Set Velocity
                                     #statPathDataValue.valueLReal := #statActualCommand.pathDataElement.cmdParameters.pathDynamics.velocity;
                                     #statModalCmdValue.valueLReal := #statModalCommand.pathDataElement.cmdParameters.pathDynamics.velocity;
                                     #statModalPrgValue.valueLReal := #statModalProgram.pathDataElement.cmdParameters.pathDynamics.velocity;

                                     // Set value with follow val from above 
                                     #tempReturnVal := "LKinLang_SetValue"(parameterValue := #tempParameterValue,
                                                                           parameterPriority := #statParameterDefinition.priorities.cmdParameters.pathDynamics.velocity,
                                                                           validCountOfParameter := #statValidCounts.cmdParameters.pathDynamics.velocity,
                                                                           parameterValueMin := #MINVAL_LREAL,
                                                                           parameterValueMax := #MAXVAL_LREAL,
                                                                           properties := #statParameterDefinition.properties,
                                                                           errorString => #statErrorString,
                                                                           parameterCounter := #statElementCounter.cmdParameters.pathDynamics.velocity,
                                                                           priorityCounter := #statActualCommand.priority.cmdParameters.pathDynamics.velocity,
                                                                           modalCMDPrio := #statModalCommand.priority.cmdParameters.pathDynamics.velocity,
                                                                           modalPRGPrio := #statModalProgram.priority.cmdParameters.pathDynamics.velocity,
                                                                           parameterCounterInLine := #statElementCounterInLine.cmdParameters.pathDynamics.velocity,
                                                                           pathDataValue := #statPathDataValue,
                                                                           modalCMDPathDataValue := #statModalCmdValue,
                                                                           modalPRGPathDataValue := #statModalPrgValue);

                                     IF #tempReturnVal = 0 THEN
                                       #statActualCommand.pathDataElement.cmdParameters.pathDynamics.velocity := #statPathDataValue.valueLReal;
                                       #statModalCommand.pathDataElement.cmdParameters.pathDynamics.velocity := #statModalCmdValue.valueLReal;
                                       #statModalProgram.pathDataElement.cmdParameters.pathDynamics.velocity := #statModalPrgValue.valueLReal;
                                     ELSE
                                       // Error
                                       #statStatus := #ERR_PARSING;
                                       #statErrorString := CONCAT(IN1 := #statErrorString, IN2 := '; Line: ');
                                       #statErrorString := CONCAT(IN1 := #statErrorString, IN2 := UDINT_TO_STRING(#statTokenizedLine.lineNo));
                                       EXIT;
                                     END_IF;
                                   END_IF;

                                   // Acceleration
                                   IF (#statParameterValid.cmdParameters.pathDynamics.acceleration AND #tempParseCounter = 1)
                                     OR (NOT #statParameterValid.cmdParameters.pathDynamics.acceleration AND #tempParseCounter = 2)
                                     AND #statParameterDefinition.priorities.cmdParameters.pathDynamics.acceleration > "LKINLANG_PRIO_UNRELEVANT"
                                   THEN

                                     // Get parameter value
                                     #tempParameterValue := #tempParsedValues.cmdParameters.pathDynamics.acceleration;

                                     // Set Velocity
                                     #statPathDataValue.valueLReal := #statActualCommand.pathDataElement.cmdParameters.pathDynamics.acceleration;
                                     #statModalCmdValue.valueLReal := #statModalCommand.pathDataElement.cmdParameters.pathDynamics.acceleration;
                                     #statModalPrgValue.valueLReal := #statModalProgram.pathDataElement.cmdParameters.pathDynamics.acceleration;

                                     // Set value with follow val from above 
                                     #tempReturnVal := "LKinLang_SetValue"(parameterValue := #tempParameterValue,
                                                                           parameterPriority := #statParameterDefinition.priorities.cmdParameters.pathDynamics.acceleration,
                                                                           validCountOfParameter := #statValidCounts.cmdParameters.pathDynamics.acceleration,
                                                                           parameterValueMin := #MINVAL_LREAL,
                                                                           parameterValueMax := #MAXVAL_LREAL,
                                                                           properties := #statParameterDefinition.properties,
                                                                           errorString => #statErrorString,
                                                                           parameterCounter := #statElementCounter.cmdParameters.pathDynamics.acceleration,
                                                                           priorityCounter := #statActualCommand.priority.cmdParameters.pathDynamics.acceleration,
                                                                           modalCMDPrio := #statModalCommand.priority.cmdParameters.pathDynamics.acceleration,
                                                                           modalPRGPrio := #statModalProgram.priority.cmdParameters.pathDynamics.acceleration,
                                                                           parameterCounterInLine := #statElementCounterInLine.cmdParameters.pathDynamics.acceleration,
                                                                           pathDataValue := #statPathDataValue,
                                                                           modalCMDPathDataValue := #statModalCmdValue,
                                                                           modalPRGPathDataValue := #statModalPrgValue);

                                     IF #tempReturnVal = 0 THEN
                                       #statActualCommand.pathDataElement.cmdParameters.pathDynamics.acceleration := #statPathDataValue.valueLReal;
                                       #statModalCommand.pathDataElement.cmdParameters.pathDynamics.acceleration := #statModalCmdValue.valueLReal;
                                       #statModalProgram.pathDataElement.cmdParameters.pathDynamics.acceleration := #statModalPrgValue.valueLReal;
                                     ELSE
                                       // Error
                                       #statStatus := #ERR_PARSING;
                                       #statErrorString := CONCAT(IN1 := #statErrorString, IN2 := '; Line: ');
                                       #statErrorString := CONCAT(IN1 := #statErrorString, IN2 := UDINT_TO_STRING(#statTokenizedLine.lineNo));
                                       EXIT;
                                     END_IF;
                                   END_IF;

                                   // Deceleration
                                   IF (#statParameterValid.cmdParameters.pathDynamics.deceleration AND #tempParseCounter = 1)
                                     OR (NOT #statParameterValid.cmdParameters.pathDynamics.deceleration AND #tempParseCounter = 2)
                                     AND #statParameterDefinition.priorities.cmdParameters.pathDynamics.deceleration > "LKINLANG_PRIO_UNRELEVANT"
                                   THEN

                                     // Get parameter value
                                     #tempParameterValue := #tempParsedValues.cmdParameters.pathDynamics.deceleration;

                                     // Set Velocity
                                     #statPathDataValue.valueLReal := #statActualCommand.pathDataElement.cmdParameters.pathDynamics.deceleration;
                                     #statModalCmdValue.valueLReal := #statModalCommand.pathDataElement.cmdParameters.pathDynamics.deceleration;
                                     #statModalPrgValue.valueLReal := #statModalProgram.pathDataElement.cmdParameters.pathDynamics.deceleration;

                                     // Set value with follow val from above 
                                     #tempReturnVal := "LKinLang_SetValue"(parameterValue := #tempParameterValue,
                                                                           parameterPriority := #statParameterDefinition.priorities.cmdParameters.pathDynamics.deceleration,
                                                                           validCountOfParameter := #statValidCounts.cmdParameters.pathDynamics.deceleration,
                                                                           parameterValueMin := #MINVAL_LREAL,
                                                                           parameterValueMax := #MAXVAL_LREAL,
                                                                           properties := #statParameterDefinition.properties,
                                                                           errorString => #statErrorString,
                                                                           parameterCounter := #statElementCounter.cmdParameters.pathDynamics.deceleration,
                                                                           priorityCounter := #statActualCommand.priority.cmdParameters.pathDynamics.deceleration,
                                                                           modalCMDPrio := #statModalCommand.priority.cmdParameters.pathDynamics.deceleration,
                                                                           modalPRGPrio := #statModalProgram.priority.cmdParameters.pathDynamics.deceleration,
                                                                           parameterCounterInLine := #statElementCounterInLine.cmdParameters.pathDynamics.deceleration,
                                                                           pathDataValue := #statPathDataValue,
                                                                           modalCMDPathDataValue := #statModalCmdValue,
                                                                           modalPRGPathDataValue := #statModalPrgValue);

                                     IF #tempReturnVal = 0 THEN
                                       #statActualCommand.pathDataElement.cmdParameters.pathDynamics.deceleration := #statPathDataValue.valueLReal;
                                       #statModalCommand.pathDataElement.cmdParameters.pathDynamics.deceleration := #statModalCmdValue.valueLReal;
                                       #statModalProgram.pathDataElement.cmdParameters.pathDynamics.deceleration := #statModalPrgValue.valueLReal;
                                     ELSE
                                       // Error
                                       #statStatus := #ERR_PARSING;
                                       #statErrorString := CONCAT(IN1 := #statErrorString, IN2 := '; Line: ');
                                       #statErrorString := CONCAT(IN1 := #statErrorString, IN2 := UDINT_TO_STRING(#statTokenizedLine.lineNo));
                                       EXIT;
                                     END_IF;
                                   END_IF;

                                   // Jerk
                                   IF (#statParameterValid.cmdParameters.pathDynamics.jerk AND #tempParseCounter = 1)
                                     OR (NOT #statParameterValid.cmdParameters.pathDynamics.jerk AND #tempParseCounter = 2)
                                     AND #statParameterDefinition.priorities.cmdParameters.pathDynamics.jerk > "LKINLANG_PRIO_UNRELEVANT"
                                   THEN

                                     // Get parameter value
                                     #tempParameterValue := #tempParsedValues.cmdParameters.pathDynamics.jerk;

                                     // Set Velocity
                                     #statPathDataValue.valueLReal := #statActualCommand.pathDataElement.cmdParameters.pathDynamics.jerk;
                                     #statModalCmdValue.valueLReal := #statModalCommand.pathDataElement.cmdParameters.pathDynamics.jerk;
                                     #statModalPrgValue.valueLReal := #statModalProgram.pathDataElement.cmdParameters.pathDynamics.jerk;

                                     // Set value with follow val from above 
                                     #tempReturnVal := "LKinLang_SetValue"(parameterValue := #tempParameterValue,
                                                                           parameterPriority := #statParameterDefinition.priorities.cmdParameters.pathDynamics.jerk,
                                                                           validCountOfParameter := #statValidCounts.cmdParameters.pathDynamics.jerk,
                                                                           parameterValueMin := #MINVAL_LREAL,
                                                                           parameterValueMax := #MAXVAL_LREAL,
                                                                           properties := #statParameterDefinition.properties,
                                                                           errorString => #statErrorString,
                                                                           parameterCounter := #statElementCounter.cmdParameters.pathDynamics.jerk,
                                                                           priorityCounter := #statActualCommand.priority.cmdParameters.pathDynamics.jerk,
                                                                           modalCMDPrio := #statModalCommand.priority.cmdParameters.pathDynamics.jerk,
                                                                           modalPRGPrio := #statModalProgram.priority.cmdParameters.pathDynamics.jerk,
                                                                           parameterCounterInLine := #statElementCounterInLine.cmdParameters.pathDynamics.jerk,
                                                                           pathDataValue := #statPathDataValue,
                                                                           modalCMDPathDataValue := #statModalCmdValue,
                                                                           modalPRGPathDataValue := #statModalPrgValue);

                                     IF #tempReturnVal = 0 THEN
                                       #statActualCommand.pathDataElement.cmdParameters.pathDynamics.jerk := #statPathDataValue.valueLReal;
                                       #statModalCommand.pathDataElement.cmdParameters.pathDynamics.jerk := #statModalCmdValue.valueLReal;
                                       #statModalProgram.pathDataElement.cmdParameters.pathDynamics.jerk := #statModalPrgValue.valueLReal;
                                     ELSE
                                       // Error
                                       #statStatus := #ERR_PARSING;
                                       #statErrorString := CONCAT(IN1 := #statErrorString, IN2 := '; Line: ');
                                       #statErrorString := CONCAT(IN1 := #statErrorString, IN2 := UDINT_TO_STRING(#statTokenizedLine.lineNo));
                                       EXIT;
                                     END_IF;
                                   END_IF;

                                 END_IF;
                               END_REGION PATH_DYNAMICS

                               REGION CIRCLE_PARAMETERS
                                 IF #tempCmdWord.%X4 THEN // Circle parameters are to be set
                                   // Aux point
                                   FOR #tempCounter := 1 TO 3 DO
                                     IF (#statParameterValid.cmdParameters.circleParameters.auxPoint[#tempCounter] AND #tempParseCounter = 1)
                                       OR (NOT #statParameterValid.cmdParameters.circleParameters.auxPoint[#tempCounter] AND #tempParseCounter = 2)
                                       AND #statParameterDefinition.priorities.cmdParameters.circleParameters.auxPoint[#tempCounter] > "LKINLANG_PRIO_UNRELEVANT"
                                     THEN

                                       // Get parameter value
                                       #tempParameterValue := #tempParsedValues.cmdParameters.circleParameters.auxPoint[#tempCounter];

                                       // Set AuxPoint
                                       #statPathDataValue.valueLReal := #statActualCommand.pathDataElement.cmdParameters.circleParameters.auxPoint[#tempCounter];
                                       #statModalCmdValue.valueLReal := #statModalCommand.pathDataElement.cmdParameters.circleParameters.auxPoint[#tempCounter];
                                       #statModalPrgValue.valueLReal := #statModalProgram.pathDataElement.cmdParameters.circleParameters.auxPoint[#tempCounter];

                                       // Set value with follow val from above 
                                       #tempReturnVal := "LKinLang_SetValue"(parameterValue := #tempParameterValue,
                                                                             parameterPriority := #statParameterDefinition.priorities.cmdParameters.circleParameters.auxPoint[#tempCounter],
                                                                             validCountOfParameter := #statValidCounts.cmdParameters.circleParameters.auxPoint[#tempCounter],
                                                                             parameterValueMin := #MINVAL_LREAL,
                                                                             parameterValueMax := #MAXVAL_LREAL,
                                                                             properties := #statParameterDefinition.properties,
                                                                             errorString => #statErrorString,
                                                                             parameterCounter := #statElementCounter.cmdParameters.circleParameters.auxPoint[#tempCounter],
                                                                             priorityCounter := #statActualCommand.priority.cmdParameters.circleParameters.auxPoint[#tempCounter],
                                                                             modalCMDPrio := #statModalCommand.priority.cmdParameters.circleParameters.auxPoint[#tempCounter],
                                                                             modalPRGPrio := #statModalProgram.priority.cmdParameters.circleParameters.auxPoint[#tempCounter],
                                                                             parameterCounterInLine := #statElementCounterInLine.cmdParameters.circleParameters.auxPoint[#tempCounter],
                                                                             pathDataValue := #statPathDataValue,
                                                                             modalCMDPathDataValue := #statModalCmdValue,
                                                                             modalPRGPathDataValue := #statModalPrgValue);

                                       IF #tempReturnVal = 0 THEN
                                         #statActualCommand.pathDataElement.cmdParameters.circleParameters.auxPoint[#tempCounter] := #statPathDataValue.valueLReal;
                                         #statModalCommand.pathDataElement.cmdParameters.circleParameters.auxPoint[#tempCounter] := #statModalCmdValue.valueLReal;
                                         #statModalProgram.pathDataElement.cmdParameters.circleParameters.auxPoint[#tempCounter] := #statModalPrgValue.valueLReal;
                                       ELSE
                                         // Error
                                         #statStatus := #ERR_PARSING;
                                         #statErrorString := CONCAT(IN1 := #statErrorString, IN2 := '; Line: ');
                                         #statErrorString := CONCAT(IN1 := #statErrorString, IN2 := UDINT_TO_STRING(#statTokenizedLine.lineNo));
                                         EXIT;
                                       END_IF;
                                     END_IF;
                                   END_FOR;

                                   // PathChoice
                                   IF (#statParameterValid.cmdParameters.circleParameters.pathChoice AND #tempParseCounter = 1)
                                     OR (NOT #statParameterValid.cmdParameters.circleParameters.pathChoice AND #tempParseCounter = 2)
                                     AND #statParameterDefinition.priorities.cmdParameters.circleParameters.pathChoice > "LKINLANG_PRIO_UNRELEVANT"
                                   THEN
                                     // Get parameter value
                                     #tempParameterValue := #tempParsedValues.cmdParameters.circleParameters.pathChoice;

                                     // Set PathChoice
                                     #statPathDataValue.valueDint := #statActualCommand.pathDataElement.cmdParameters.circleParameters.pathChoice;
                                     #statModalCmdValue.valueDint := #statModalCommand.pathDataElement.cmdParameters.circleParameters.pathChoice;
                                     #statModalPrgValue.valueDint := #statModalProgram.pathDataElement.cmdParameters.circleParameters.pathChoice;

                                     // Set value with follow val from above 
                                     #tempReturnVal := "LKinLang_SetValue"(parameterValue := #tempParameterValue,
                                                                           parameterPriority := #statParameterDefinition.priorities.cmdParameters.circleParameters.pathChoice,
                                                                           validCountOfParameter := #statValidCounts.cmdParameters.circleParameters.pathChoice,
                                                                           parameterValueMin := 0,
                                                                           parameterValueMax := 3,
                                                                           properties := #statParameterDefinition.properties,
                                                                           errorString => #statErrorString,
                                                                           parameterCounter := #statElementCounter.cmdParameters.circleParameters.pathChoice,
                                                                           priorityCounter := #statActualCommand.priority.cmdParameters.circleParameters.pathChoice,
                                                                           modalCMDPrio := #statModalCommand.priority.cmdParameters.circleParameters.pathChoice,
                                                                           modalPRGPrio := #statModalProgram.priority.cmdParameters.circleParameters.pathChoice,
                                                                           parameterCounterInLine := #statElementCounterInLine.cmdParameters.circleParameters.pathChoice,
                                                                           pathDataValue := #statPathDataValue,
                                                                           modalCMDPathDataValue := #statModalCmdValue,
                                                                           modalPRGPathDataValue := #statModalPrgValue);

                                     IF #tempReturnVal = 0 THEN
                                       #statActualCommand.pathDataElement.cmdParameters.circleParameters.pathChoice := #statPathDataValue.valueDint;
                                       #statModalCommand.pathDataElement.cmdParameters.circleParameters.pathChoice := #statModalCmdValue.valueDint;
                                       #statModalProgram.pathDataElement.cmdParameters.circleParameters.pathChoice := #statModalPrgValue.valueDint;
                                     ELSE
                                       // Error
                                       #statStatus := #ERR_PARSING;
                                       #statErrorString := CONCAT(IN1 := #statErrorString, IN2 := '; Line: ');
                                       #statErrorString := CONCAT(IN1 := #statErrorString, IN2 := UDINT_TO_STRING(#statTokenizedLine.lineNo));
                                       EXIT;
                                     END_IF;
                                   END_IF;


                                   // CircMode
                                   IF (#statParameterValid.cmdParameters.circleParameters.circMode AND #tempParseCounter = 1)
                                     OR (NOT #statParameterValid.cmdParameters.circleParameters.circMode AND #tempParseCounter = 2)
                                     AND #statParameterDefinition.priorities.cmdParameters.circleParameters.circMode > "LKINLANG_PRIO_UNRELEVANT"
                                   THEN
                                     // Get parameter value
                                     #tempParameterValue := #tempParsedValues.cmdParameters.circleParameters.circMode;

                                     // Set CircMode
                                     #statPathDataValue.valueDint := #statActualCommand.pathDataElement.cmdParameters.circleParameters.circMode;
                                     #statModalCmdValue.valueDint := #statModalCommand.pathDataElement.cmdParameters.circleParameters.circMode;
                                     #statModalPrgValue.valueDint := #statModalProgram.pathDataElement.cmdParameters.circleParameters.circMode;

                                     // Set value with follow val from above 
                                     #tempReturnVal := "LKinLang_SetValue"(parameterValue := #tempParameterValue,
                                                                           parameterPriority := #statParameterDefinition.priorities.cmdParameters.circleParameters.circMode,
                                                                           validCountOfParameter := #statValidCounts.cmdParameters.circleParameters.circMode,
                                                                           parameterValueMin := 0,
                                                                           parameterValueMax := 2,
                                                                           properties := #statParameterDefinition.properties,
                                                                           errorString => #statErrorString,
                                                                           parameterCounter := #statElementCounter.cmdParameters.circleParameters.circMode,
                                                                           priorityCounter := #statActualCommand.priority.cmdParameters.circleParameters.circMode,
                                                                           modalCMDPrio := #statModalCommand.priority.cmdParameters.circleParameters.circMode,
                                                                           modalPRGPrio := #statModalProgram.priority.cmdParameters.circleParameters.circMode,
                                                                           parameterCounterInLine := #statElementCounterInLine.cmdParameters.circleParameters.circMode,
                                                                           pathDataValue := #statPathDataValue,
                                                                           modalCMDPathDataValue := #statModalCmdValue,
                                                                           modalPRGPathDataValue := #statModalPrgValue);

                                     IF #tempReturnVal = 0 THEN
                                       #statActualCommand.pathDataElement.cmdParameters.circleParameters.circMode := #statPathDataValue.valueDint;
                                       #statModalCommand.pathDataElement.cmdParameters.circleParameters.circMode := #statModalCmdValue.valueDint;
                                       #statModalProgram.pathDataElement.cmdParameters.circleParameters.circMode := #statModalPrgValue.valueDint;
                                     ELSE
                                       // Error
                                       #statStatus := #ERR_PARSING;
                                       #statErrorString := CONCAT(IN1 := #statErrorString, IN2 := '; Line: ');
                                       #statErrorString := CONCAT(IN1 := #statErrorString, IN2 := UDINT_TO_STRING(#statTokenizedLine.lineNo));
                                       EXIT;
                                     END_IF;
                                   END_IF;


                                   // CirclePlane
                                   IF (#statParameterValid.cmdParameters.circleParameters.circlePlane AND #tempParseCounter = 1)
                                     OR (NOT #statParameterValid.cmdParameters.circleParameters.circlePlane AND #tempParseCounter = 2)
                                     AND #statParameterDefinition.priorities.cmdParameters.circleParameters.circlePlane > "LKINLANG_PRIO_UNRELEVANT"
                                   THEN
                                     // Get parameter value
                                     #tempParameterValue := #tempParsedValues.cmdParameters.circleParameters.circlePlane;

                                     // Set CirclePlane
                                     #statPathDataValue.valueDint := #statActualCommand.pathDataElement.cmdParameters.circleParameters.circlePlane;
                                     #statModalCmdValue.valueDint := #statModalCommand.pathDataElement.cmdParameters.circleParameters.circlePlane;
                                     #statModalPrgValue.valueDint := #statModalProgram.pathDataElement.cmdParameters.circleParameters.circlePlane;

                                     // Set value with follow val from above 
                                     #tempReturnVal := "LKinLang_SetValue"(parameterValue := #tempParameterValue,
                                                                           parameterPriority := #statParameterDefinition.priorities.cmdParameters.circleParameters.circlePlane,
                                                                           validCountOfParameter := #statValidCounts.cmdParameters.circleParameters.circlePlane,
                                                                           parameterValueMin := 0,
                                                                           parameterValueMax := 2,
                                                                           properties := #statParameterDefinition.properties,
                                                                           errorString => #statErrorString,
                                                                           parameterCounter := #statElementCounter.cmdParameters.circleParameters.circlePlane,
                                                                           priorityCounter := #statActualCommand.priority.cmdParameters.circleParameters.circlePlane,
                                                                           modalCMDPrio := #statModalCommand.priority.cmdParameters.circleParameters.circlePlane,
                                                                           modalPRGPrio := #statModalProgram.priority.cmdParameters.circleParameters.circlePlane,
                                                                           parameterCounterInLine := #statElementCounterInLine.cmdParameters.circleParameters.circlePlane,
                                                                           pathDataValue := #statPathDataValue,
                                                                           modalCMDPathDataValue := #statModalCmdValue,
                                                                           modalPRGPathDataValue := #statModalPrgValue);

                                     IF #tempReturnVal = 0 THEN
                                       #statActualCommand.pathDataElement.cmdParameters.circleParameters.circlePlane := #statPathDataValue.valueDint;
                                       #statModalCommand.pathDataElement.cmdParameters.circleParameters.circlePlane := #statModalCmdValue.valueDint;
                                       #statModalProgram.pathDataElement.cmdParameters.circleParameters.circlePlane := #statModalPrgValue.valueDint;
                                     ELSE
                                       // Error
                                       #statStatus := #ERR_PARSING;
                                       #statErrorString := CONCAT(IN1 := #statErrorString, IN2 := '; Line: ');
                                       #statErrorString := CONCAT(IN1 := #statErrorString, IN2 := UDINT_TO_STRING(#statTokenizedLine.lineNo));
                                       EXIT;
                                     END_IF;
                                   END_IF;


